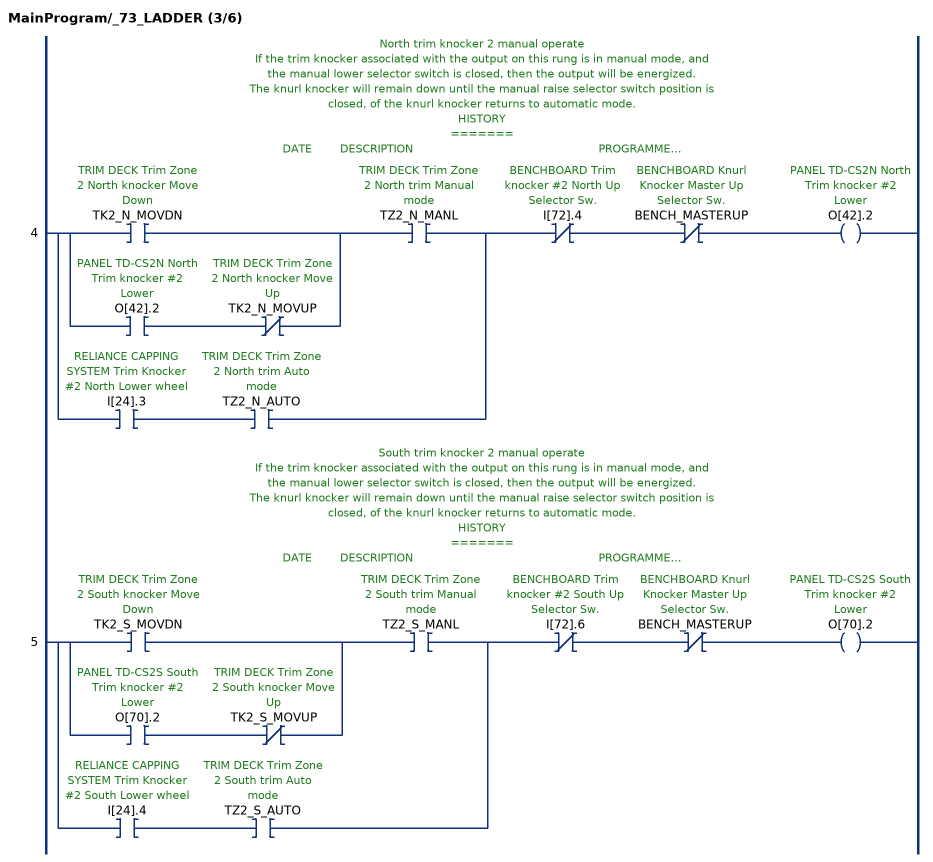
   // North trim knocker 2 manual operate
   // If the trim knocker associated with the output on this rung is in manual mode, and
   // the manual lower selector switch is closed, then the output will be energized.
   // The knurl knocker will remain down until the manual raise selector switch position is
   // closed, of the knurl knocker returns to automatic mode.
   // HISTORY
   // =======
   // DATE        DESCRIPTION                                                     PROGRAMMER
   // ====        ===========                                                     ==========
   // 2/29/96     Entered rung as designed                                        WAS
   // 3/1/96      Added these comments                                            WAS
   4: [[XIC(TK2_N_MOVDN) ,XIC(O[42].2) XIO(TK2_N_MOVUP) ] XIC(TZ2_N_MANL) ,XIC(I[24].3) XIC(TZ2_N_AUTO) ]XIO(I[72].4)XIO(BENCH_MASTERUP)OTE(O[42].2);
   // South trim knocker 2 manual operate
   // If the trim knocker associated with the output on this rung is in manual mode, and
   // the manual lower selector switch is closed, then the output will be energized.
   // The knurl knocker will remain down until the manual raise selector switch position is
   // closed, of the knurl knocker returns to automatic mode.
   // HISTORY
   // =======
   // DATE        DESCRIPTION                                                     PROGRAMMER
   // ====        ===========                                                     ==========
   // 2/29/96     Entered rung as designed                                        WAS
   // 3/1/96      Added these comments                                            WAS
   5: [[XIC(TK2_S_MOVDN) ,XIC(O[70].2) XIO(TK2_S_MOVUP) ] XIC(TZ2_S_MANL) ,XIC(I[24].4) XIC(TZ2_S_AUTO) ]XIO(I[72].6)XIO(BENCH_MASTERUP)OTE(O[70].2);
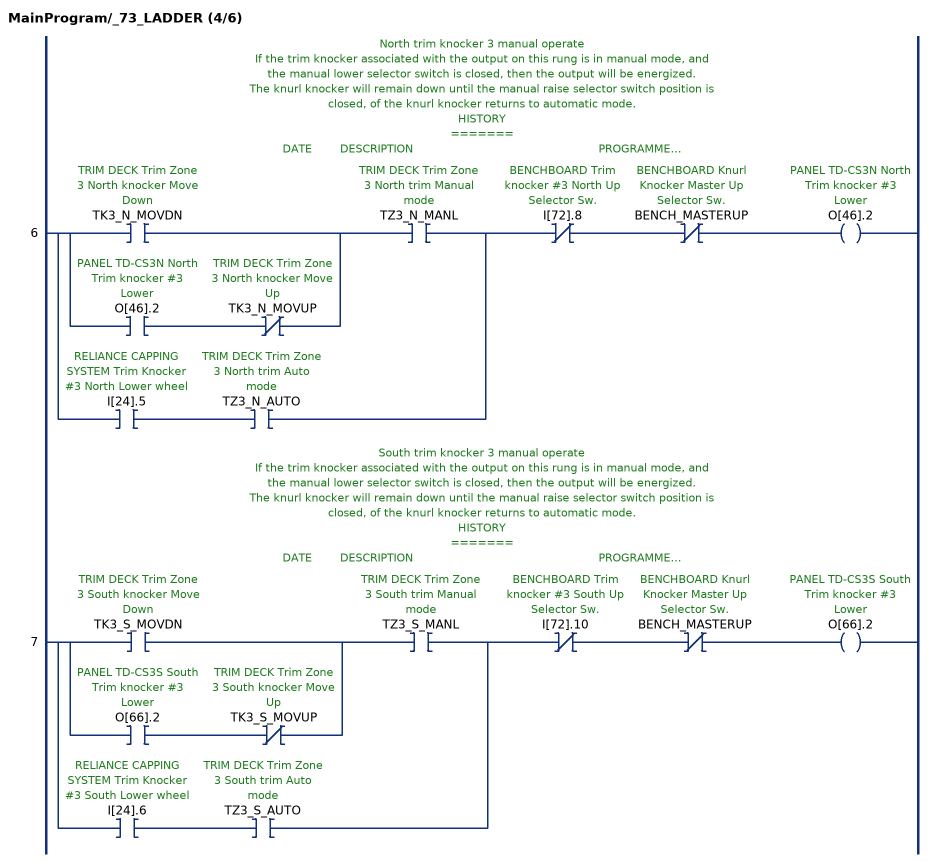
   // North trim knocker 3 manual operate
   // If the trim knocker associated with the output on this rung is in manual mode, and
   // the manual lower selector switch is closed, then the output will be energized.
   // The knurl knocker will remain down until the manual raise selector switch position is
   // closed, of the knurl knocker returns to automatic mode.
   // HISTORY
   // =======
   // DATE        DESCRIPTION                                                     PROGRAMMER
   // ====        ===========                                                     ==========
   // 2/29/96     Entered rung as designed                                        WAS
   // 3/1/96      Added these comments                                            WAS
   6: [[XIC(TK3_N_MOVDN) ,XIC(O[46].2) XIO(TK3_N_MOVUP) ] XIC(TZ3_N_MANL) ,XIC(I[24].5) XIC(TZ3_N_AUTO) ]XIO(I[72].8)XIO(BENCH_MASTERUP)OTE(O[46].2);
   // South trim knocker 3 manual operate
   // If the trim knocker associated with the output on this rung is in manual mode, and
   // the manual lower selector switch is closed, then the output will be energized.
   // The knurl knocker will remain down until the manual raise selector switch position is
   // closed, of the knurl knocker returns to automatic mode.
   // HISTORY
   // =======
   // DATE        DESCRIPTION                                                     PROGRAMMER
   // ====        ===========                                                     ==========
   // 2/29/96     Entered rung as designed                                        WAS
   // 3/1/96      Added these comments                                            WAS
   7: [[XIC(TK3_S_MOVDN) ,XIC(O[66].2) XIO(TK3_S_MOVUP) ] XIC(TZ3_S_MANL) ,XIC(I[24].6) XIC(TZ3_S_AUTO) ]XIO(I[72].10)XIO(BENCH_MASTERUP)OTE(O[66].2);
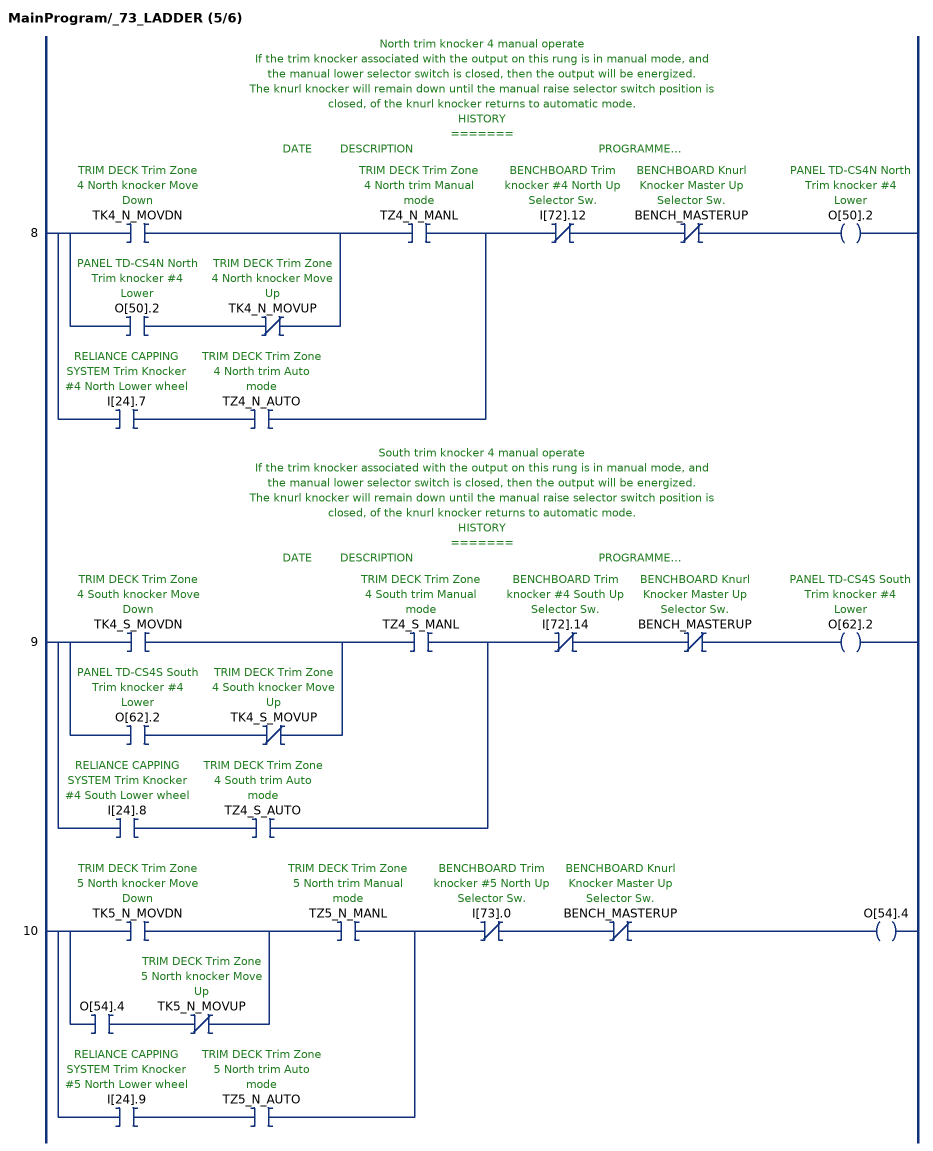
   // North trim knocker 4 manual operate
   // If the trim knocker associated with the output on this rung is in manual mode, and
   // the manual lower selector switch is closed, then the output will be energized.
   // The knurl knocker will remain down until the manual raise selector switch position is
   // closed, of the knurl knocker returns to automatic mode.
   // HISTORY
   // =======
   // DATE        DESCRIPTION                                                     PROGRAMMER
   // ====        ===========                                                     ==========
   // 2/29/96     Entered rung as designed                                        WAS
   // 3/1/96      Added these comments                                            WAS
   8: [[XIC(TK4_N_MOVDN) ,XIC(O[50].2) XIO(TK4_N_MOVUP) ] XIC(TZ4_N_MANL) ,XIC(I[24].7) XIC(TZ4_N_AUTO) ]XIO(I[72].12)XIO(BENCH_MASTERUP)OTE(O[50].2);
   // South trim knocker 4 manual operate
   // If the trim knocker associated with the output on this rung is in manual mode, and
   // the manual lower selector switch is closed, then the output will be energized.
   // The knurl knocker will remain down until the manual raise selector switch position is
   // closed, of the knurl knocker returns to automatic mode.
   // HISTORY
   // =======
   // DATE        DESCRIPTION                                                     PROGRAMMER
   // ====        ===========                                                     ==========
   // 2/29/96     Entered rung as designed                                        WAS
   // 3/1/96      Added these comments                                            WAS
   9: [[XIC(TK4_S_MOVDN) ,XIC(O[62].2) XIO(TK4_S_MOVUP) ] XIC(TZ4_S_MANL) ,XIC(I[24].8) XIC(TZ4_S_AUTO) ]XIO(I[72].14)XIO(BENCH_MASTERUP)OTE(O[62].2);
   10: [[XIC(TK5_N_MOVDN) ,XIC(O[54].4) XIO(TK5_N_MOVUP) ] XIC(TZ5_N_MANL) ,XIC(I[24].9) XIC(TZ5_N_AUTO) ]XIO(I[73].0)XIO(BENCH_MASTERUP)OTE(O[54].4);
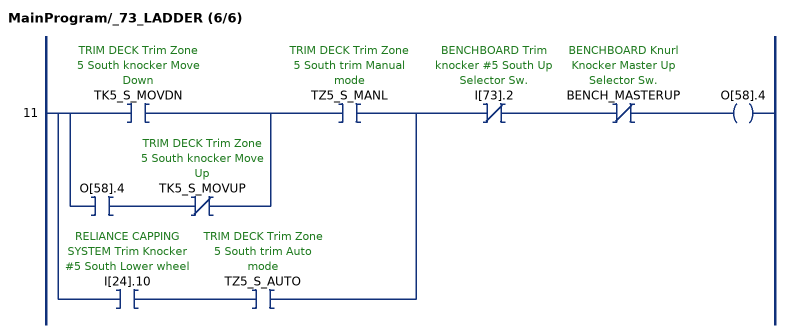
   11: [[XIC(TK5_S_MOVDN) ,XIC(O[58].4) XIO(TK5_S_MOVUP) ] XIC(TZ5_S_MANL) ,XIC(I[24].10) XIC(TZ5_S_AUTO) ]XIO(I[73].2)XIO(BENCH_MASTERUP)OTE(O[58].4);
END_ROUTINE

ROUTINE _74_LADDER   (* ladder *)
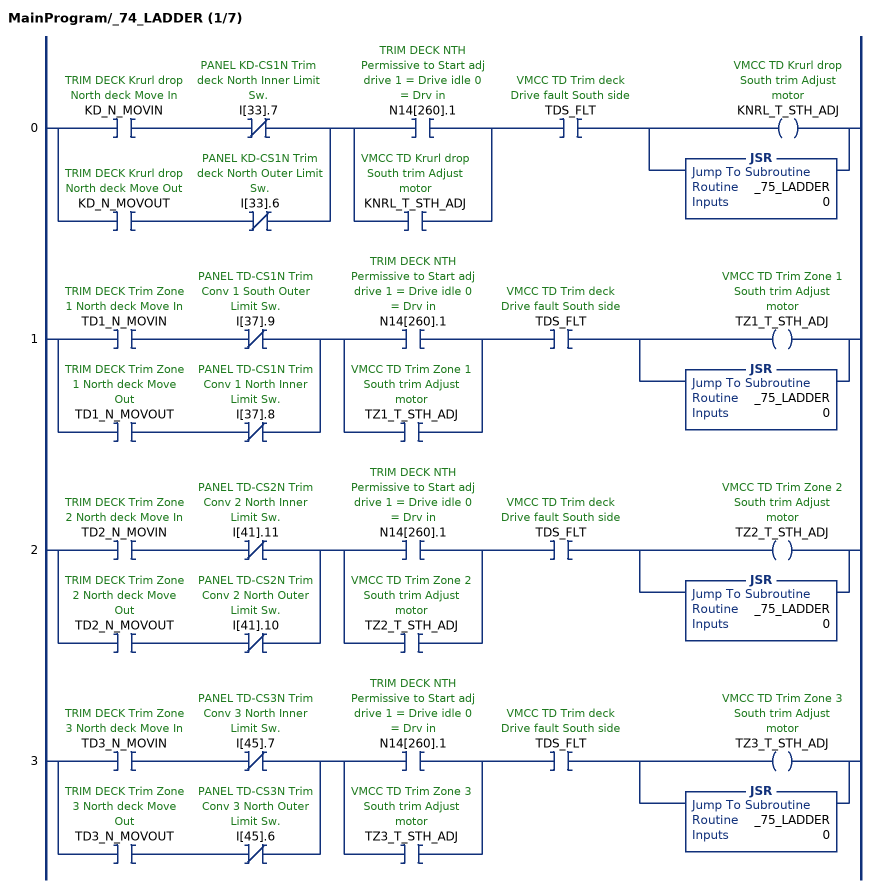
   0: [XIC(KD_N_MOVIN) XIO(I[33].7) ,XIC(KD_N_MOVOUT) XIO(I[33].6) ][XIC(N14[260].1) ,XIC(KNRL_T_STH_ADJ) ]XIC(TDS_FLT)[OTE(KNRL_T_STH_ADJ) ,JSR(_75_LADDER,0) ];
   1: [XIC(TD1_N_MOVIN) XIO(I[37].9) ,XIC(TD1_N_MOVOUT) XIO(I[37].8) ][XIC(N14[260].1) ,XIC(TZ1_T_STH_ADJ) ]XIC(TDS_FLT)[OTE(TZ1_T_STH_ADJ) ,JSR(_75_LADDER,0) ];
   2: [XIC(TD2_N_MOVIN) XIO(I[41].11) ,XIC(TD2_N_MOVOUT) XIO(I[41].10) ][XIC(N14[260].1) ,XIC(TZ2_T_STH_ADJ) ]XIC(TDS_FLT)[OTE(TZ2_T_STH_ADJ) ,JSR(_75_LADDER,0) ];
   3: [XIC(TD3_N_MOVIN) XIO(I[45].7) ,XIC(TD3_N_MOVOUT) XIO(I[45].6) ][XIC(N14[260].1) ,XIC(TZ3_T_STH_ADJ) ]XIC(TDS_FLT)[OTE(TZ3_T_STH_ADJ) ,JSR(_75_LADDER,0) ];
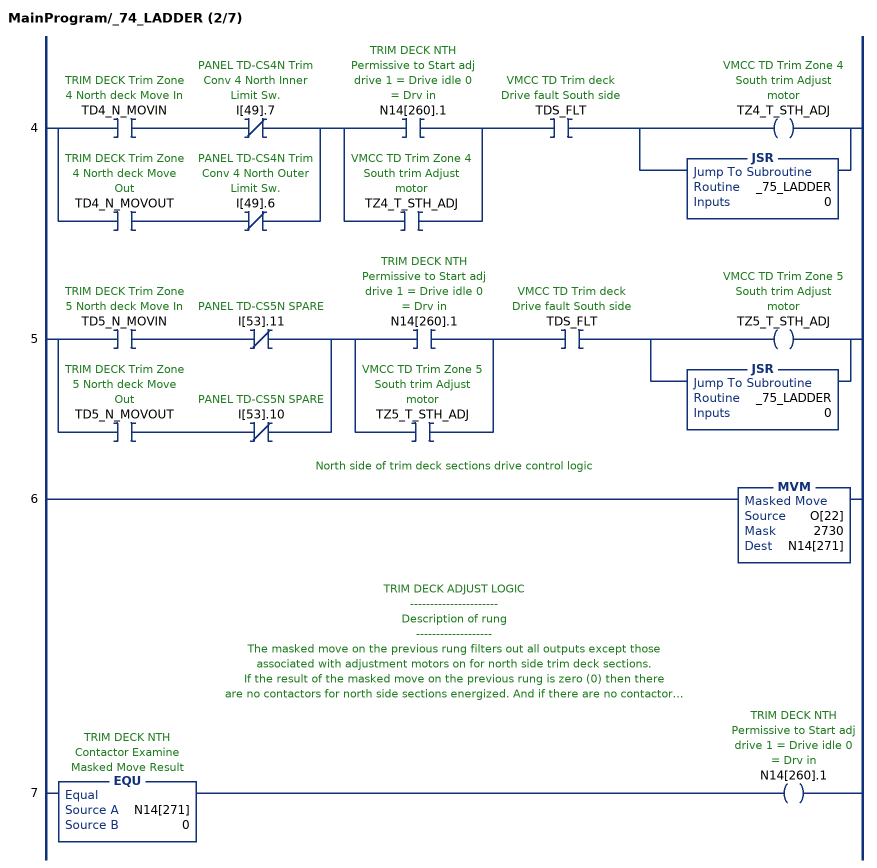
   4: [XIC(TD4_N_MOVIN) XIO(I[49].7) ,XIC(TD4_N_MOVOUT) XIO(I[49].6) ][XIC(N14[260].1) ,XIC(TZ4_T_STH_ADJ) ]XIC(TDS_FLT)[OTE(TZ4_T_STH_ADJ) ,JSR(_75_LADDER,0) ];
   5: [XIC(TD5_N_MOVIN) XIO(I[53].11) ,XIC(TD5_N_MOVOUT) XIO(I[53].10) ][XIC(N14[260].1) ,XIC(TZ5_T_STH_ADJ) ]XIC(TDS_FLT)[OTE(TZ5_T_STH_ADJ) ,JSR(_75_LADDER,0) ];
   // North side of trim deck sections drive control logic
   6: MVM(O[22],2730,N14[271]);
   // TRIM DECK ADJUST LOGIC
   // ----------------------
   // Description of rung
   // -------------------
   // The masked move on the previous rung filters out all outputs except those
   // associated with adjustment motors on for north side trim deck sections.
   // If the result of the masked move on the previous rung is zero (0) then there
   // are no contactors for north side sections energized. And if there are no contactors
   // for north side sections energized, then any north section may be energized.
   // As soon as the contactor for any section energizes, the result of the mased move on the
   // HISTORY
   // =======
   // DATE        DESCRIPTION                                                       PROGRAMMER
   // ====        ===========                                                       ==========
   // 2/29/96     Entered rung as designed                                          WAS
   // 3/1/96      Entered comment                                                   WAS
   7: EQU(N14[271],0)OTE(N14[260].1);
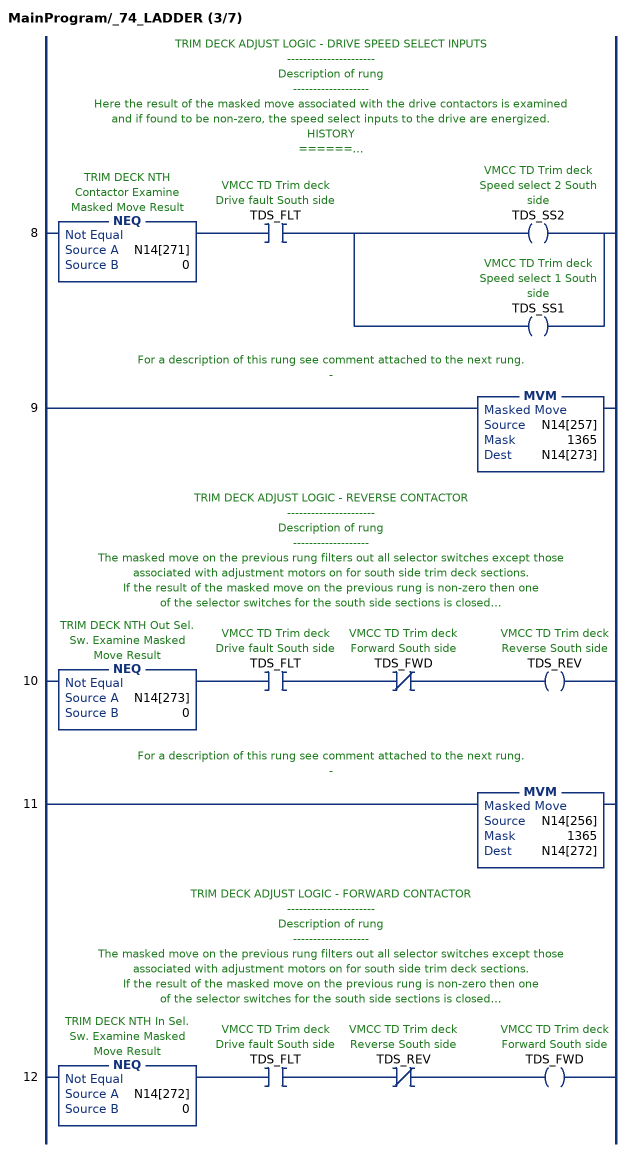
   // TRIM DECK ADJUST LOGIC - DRIVE SPEED SELECT INPUTS
   // ----------------------
   // Description of rung
   // -------------------
   // Here the result of the masked move associated with the drive contactors is examined
   // and if found to be non-zero, the speed select inputs to the drive are energized.
   // HISTORY
   // =======
   // DATE        DESCRIPTION                                                       PROGRAMMER
   // ====        ===========                                                       ==========
   // 2/29/96     Entered rung as designed                                          WAS
   // 3/1/96      Entered comment                                                   WAS
   8: NEQ(N14[271],0)XIC(TDS_FLT)[OTE(TDS_SS2) ,OTE(TDS_SS1) ];
   // For a description of this rung see comment attached to the next rung.
   //                                                                                                          -
   9: MVM(N14[257],1365,N14[273]);
   // TRIM DECK ADJUST LOGIC - REVERSE CONTACTOR
   // ----------------------
   // Description of rung
   // -------------------
   // The masked move on the previous rung filters out all selector switches except those
   // associated with adjustment motors on for south side trim deck sections.
   // If the result of the masked move on the previous rung is non-zero then one
   // of the selector switches for the south side sections is closed.
   // The selector switches examined on this rung are for outward movement, away from the
   // center of the conveyors. Any movement in this direction is accomplished by operating the
   // adjust motor in reverse. Hence, if any of the out selector switches is made, then
   // the reverse drive inpu should be energized.
   // HISTORY
   // =======
   // DATE        DESCRIPTION                                                       PROGRAMMER
   // ====        ===========                                                       ==========
   // 2/29/96     Entered rung as designed                                          WAS
   // 3/1/96      Entered comment                                                   WAS
   10: NEQ(N14[273],0)XIC(TDS_FLT)XIO(TDS_FWD)OTE(TDS_REV);
   // For a description of this rung see comment attached to the next rung.
   //                                                                                                          -
   11: MVM(N14[256],1365,N14[272]);
   // TRIM DECK ADJUST LOGIC - FORWARD CONTACTOR
   // ----------------------
   // Description of rung
   // -------------------
   // The masked move on the previous rung filters out all selector switches except those
   // associated with adjustment motors on for south side trim deck sections.
   // If the result of the masked move on the previous rung is non-zero then one
   // of the selector switches for the south side sections is closed.
   // The selector switches examined on this rung are for INWARD movement, toward the
   // center of the conveyors. Any movement in this direction is accomplished by operating the
   // adjust motor in the forward direction. Hence, if any of the out selector switches is made, then
   // the forward drive input should be energized.
   // HISTORY
   // =======
   // DATE        DESCRIPTION                                                       PROGRAMMER
   // ====        ===========                                                       ==========
   // 2/29/96     Entered rung as designed                                          WAS
   // 3/1/96      Entered comment                                                   WAS
   12: NEQ(N14[272],0)XIC(TDS_FLT)XIO(TDS_REV)OTE(TDS_FWD);
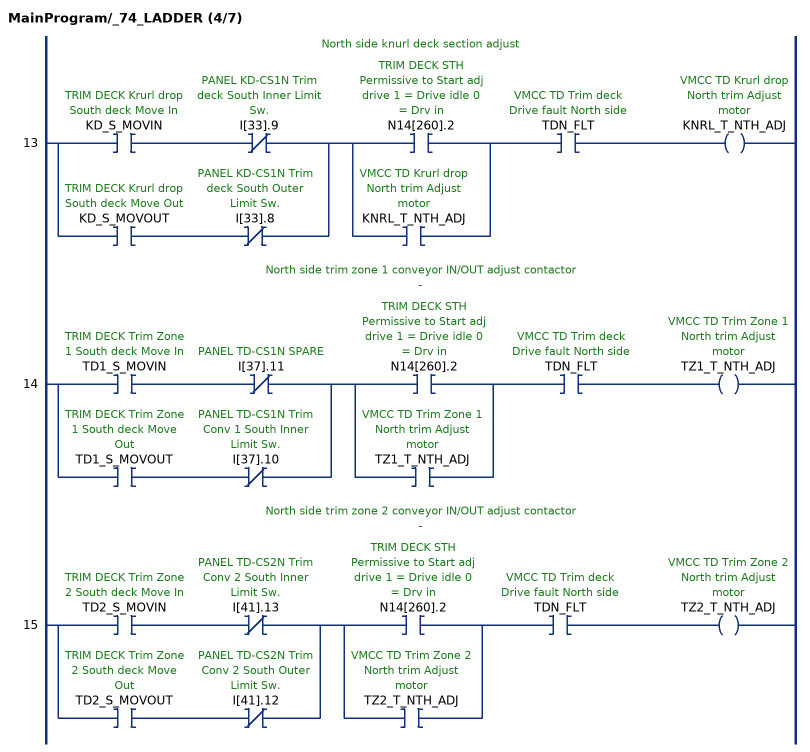
   // North side knurl deck section adjust
   13: [XIC(KD_S_MOVIN) XIO(I[33].9) ,XIC(KD_S_MOVOUT) XIO(I[33].8) ][XIC(N14[260].2) ,XIC(KNRL_T_NTH_ADJ) ]XIC(TDN_FLT)OTE(KNRL_T_NTH_ADJ);
   // North side trim zone 1 conveyor IN/OUT adjust contactor
   //                                                                                                 -
   14: [XIC(TD1_S_MOVIN) XIO(I[37].11) ,XIC(TD1_S_MOVOUT) XIO(I[37].10) ][XIC(N14[260].2) ,XIC(TZ1_T_NTH_ADJ) ]XIC(TDN_FLT)OTE(TZ1_T_NTH_ADJ);
   // North side trim zone 2 conveyor IN/OUT adjust contactor
   //                                                                                                 -
   15: [XIC(TD2_S_MOVIN) XIO(I[41].13) ,XIC(TD2_S_MOVOUT) XIO(I[41].12) ][XIC(N14[260].2) ,XIC(TZ2_T_NTH_ADJ) ]XIC(TDN_FLT)OTE(TZ2_T_NTH_ADJ);
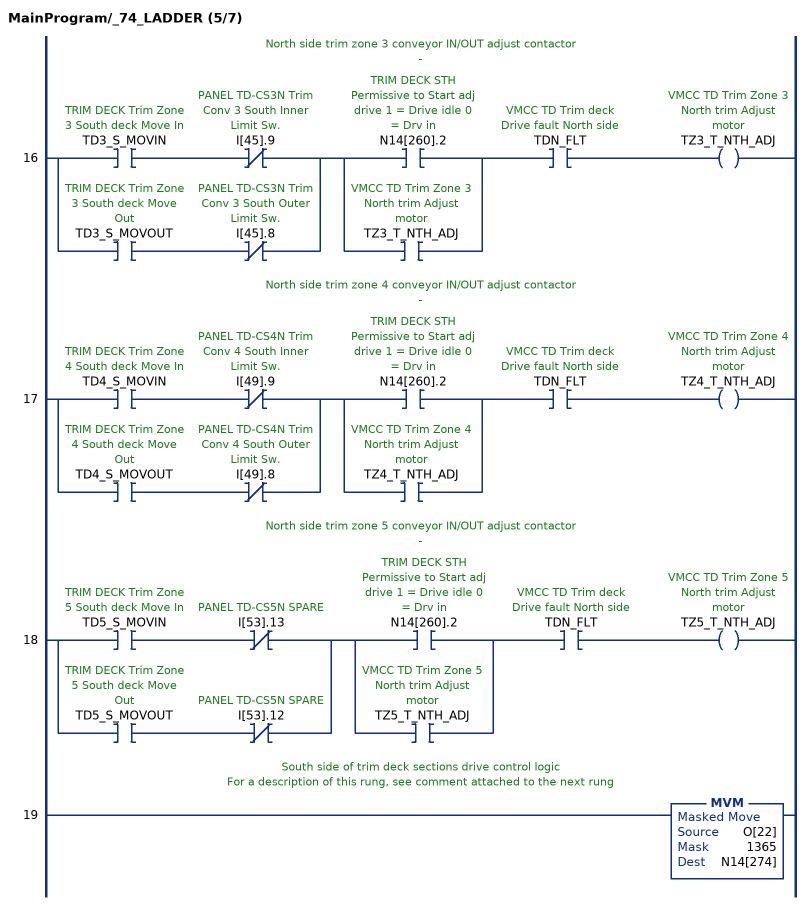
   // North side trim zone 3 conveyor IN/OUT adjust contactor
   //                                                                                                 -
   16: [XIC(TD3_S_MOVIN) XIO(I[45].9) ,XIC(TD3_S_MOVOUT) XIO(I[45].8) ][XIC(N14[260].2) ,XIC(TZ3_T_NTH_ADJ) ]XIC(TDN_FLT)OTE(TZ3_T_NTH_ADJ);
   // North side trim zone 4 conveyor IN/OUT adjust contactor
   //                                                                                                 -
   17: [XIC(TD4_S_MOVIN) XIO(I[49].9) ,XIC(TD4_S_MOVOUT) XIO(I[49].8) ][XIC(N14[260].2) ,XIC(TZ4_T_NTH_ADJ) ]XIC(TDN_FLT)OTE(TZ4_T_NTH_ADJ);
   // North side trim zone 5 conveyor IN/OUT adjust contactor
   //                                                                                                 -
   18: [XIC(TD5_S_MOVIN) XIO(I[53].13) ,XIC(TD5_S_MOVOUT) XIO(I[53].12) ][XIC(N14[260].2) ,XIC(TZ5_T_NTH_ADJ) ]XIC(TDN_FLT)OTE(TZ5_T_NTH_ADJ);
   // South side of trim deck sections drive control logic
   // For a description of this rung, see comment attached to the next rung
   19: MVM(O[22],1365,N14[274]);
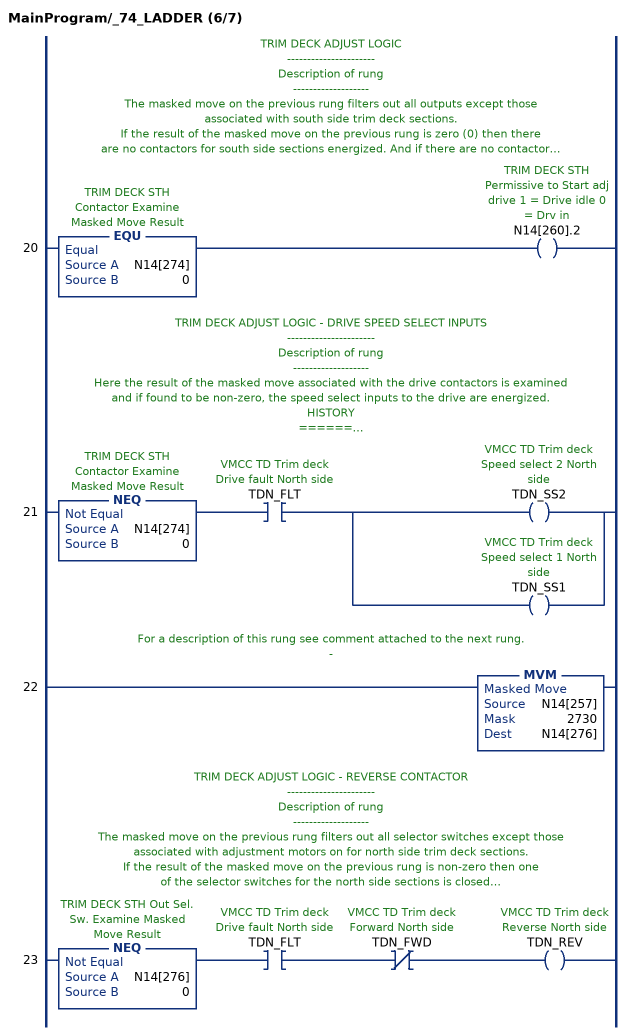
   // TRIM DECK ADJUST LOGIC
   // ----------------------
   // Description of rung
   // -------------------
   // The masked move on the previous rung filters out all outputs except those
   // associated with south side trim deck sections.
   // If the result of the masked move on the previous rung is zero (0) then there
   // are no contactors for south side sections energized. And if there are no contactors
   // for south side sections energized, then any north section may be energized.
   // As soon as the contactor for any section energizes, the result of the mased move on the
   // HISTORY
   // =======
   // DATE        DESCRIPTION                                                       PROGRAMMER
   // ====        ===========                                                       ==========
   // 2/29/96     Entered rung as designed                                          WAS
   // 3/1/96      Entered comment                                                   WAS
   // previous rung becomes non-zero, prohibiting any other sections from energizing.
   20: EQU(N14[274],0)OTE(N14[260].2);
   // TRIM DECK ADJUST LOGIC - DRIVE SPEED SELECT INPUTS
   // ----------------------
   // Description of rung
   // -------------------
   // Here the result of the masked move associated with the drive contactors is examined
   // and if found to be non-zero, the speed select inputs to the drive are energized.
   // HISTORY
   // =======
   // DATE        DESCRIPTION                                                       PROGRAMMER
   // ====        ===========                                                       ==========
   // 2/29/96     Entered rung as designed                                          WAS
   // 3/1/96      Entered comment                                                   WAS
   21: NEQ(N14[274],0)XIC(TDN_FLT)[OTE(TDN_SS2) ,OTE(TDN_SS1) ];
   // For a description of this rung see comment attached to the next rung.
   //                                                                                                          -
   22: MVM(N14[257],2730,N14[276]);
   // TRIM DECK ADJUST LOGIC - REVERSE CONTACTOR
   // ----------------------
   // Description of rung
   // -------------------
   // The masked move on the previous rung filters out all selector switches except those
   // associated with adjustment motors on for north side trim deck sections.
   // If the result of the masked move on the previous rung is non-zero then one
   // of the selector switches for the north side sections is closed.
   // The selector switches examined on this rung are for outward movement, away from the
   // center of the conveyors. Any movement in this direction is accomplished by operating the
   // adjust motor in reverse. Hence, if any of the out selector switches is made, then
   // the reverse drive inpu should be energized.
   // HISTORY
   // =======
   // DATE        DESCRIPTION                                                       PROGRAMMER
   // ====        ===========                                                       ==========
   // 2/29/96     Entered rung as designed                                          WAS
   // 3/1/96      Entered comment                                                   WAS
   23: NEQ(N14[276],0)XIC(TDN_FLT)XIO(TDN_FWD)OTE(TDN_REV);
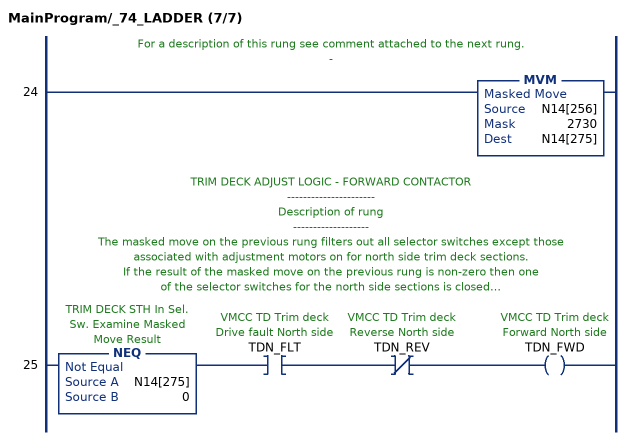
   // For a description of this rung see comment attached to the next rung.
   //                                                                                                          -
   24: MVM(N14[256],2730,N14[275]);
   // TRIM DECK ADJUST LOGIC - FORWARD CONTACTOR
   // ----------------------
   // Description of rung
   // -------------------
   // The masked move on the previous rung filters out all selector switches except those
   // associated with adjustment motors on for north side trim deck sections.
   // If the result of the masked move on the previous rung is non-zero then one
   // of the selector switches for the north side sections is closed.
   // The selector switches examined on this rung are for INWARD movement, toward the
   // center of the conveyors. Any movement in this direction is accomplished by operating the
   // adjust motor in the forward direction. Hence, if any of the out selector switches is made, then
   // the forward drive input should be energized.
   // HISTORY
   // =======
   // DATE        DESCRIPTION                                                       PROGRAMMER
   // ====        ===========                                                       ==========
   // 2/29/96     Entered rung as designed                                          WAS
   // 3/1/96      Entered comment                                                   WAS
   25: NEQ(N14[275],0)XIC(TDN_FLT)XIO(TDN_REV)OTE(TDN_FWD);
END_ROUTINE
